HMI tags "DB_SDC_ERROR_STAT_EMS057"
   "DB_SDC_ERRORS_STAT_ER_AKT[57].ER_TRIGER" : Word = PLC DB_SDC_ERRORS_STAT.ER_AKT[57].ER_TRIGER AT %DB3724.DBW31716, 1 s
   "DB_SDC_ERRORS_STAT_ER_AKT[57].ER_STAT[1].DRIVE_POS" : DInt = PLC DB_SDC_ERRORS_STAT.ER_AKT[57].ER_STAT[1].DRIVE_POS AT %DB3724.DBD31722, 1 s
   "DB_SDC_ERRORS_STAT_ER_AKT[57].ER_STAT[1].ERROR" : Int = PLC DB_SDC_ERRORS_STAT.ER_AKT[57].ER_STAT[1].ERROR AT %DB3724.DBW31728, 1 s
   "DB_SDC_ERRORS_STAT_ER_AKT[57].ER_STAT[2].DRIVE_POS" : DInt = PLC DB_SDC_ERRORS_STAT.ER_AKT[57].ER_STAT[2].DRIVE_POS AT %DB3724.DBD31738, 1 s
   "DB_SDC_ERRORS_STAT_ER_AKT[57].ER_STAT[2].ERROR" : Int = PLC DB_SDC_ERRORS_STAT.ER_AKT[57].ER_STAT[2].ERROR AT %DB3724.DBW31744, 1 s
   "DB_SDC_ERRORS_STAT_ER_AKT[57].ER_STAT[3].DRIVE_POS" : DInt = PLC DB_SDC_ERRORS_STAT.ER_AKT[57].ER_STAT[3].DRIVE_POS AT %DB3724.DBD31754, 1 s
   "DB_SDC_ERRORS_STAT_ER_AKT[57].ER_STAT[3].ERROR" : Int = PLC DB_SDC_ERRORS_STAT.ER_AKT[57].ER_STAT[3].ERROR AT %DB3724.DBW31760, 1 s
   "DB_SDC_ERRORS_STAT_ER_AKT[57].ER_STAT[4].DRIVE_POS" : DInt = PLC DB_SDC_ERRORS_STAT.ER_AKT[57].ER_STAT[4].DRIVE_POS AT %DB3724.DBD31770, 1 s
   "DB_SDC_ERRORS_STAT_ER_AKT[57].ER_STAT[4].ERROR" : Int = PLC DB_SDC_ERRORS_STAT.ER_AKT[57].ER_STAT[4].ERROR AT %DB3724.DBW31776, 1 s

HMI tags "DB_SDC_ERROR_STAT_EMS058"
   "DB_SDC_ERRORS_STAT_ER_AKT[58].ER_TRIGER" : Word = PLC DB_SDC_ERRORS_STAT.ER_AKT[58].ER_TRIGER AT %DB3724.DBW31782, 1 s
   "DB_SDC_ERRORS_STAT_ER_AKT[58].ER_STAT[1].DRIVE_POS" : DInt = PLC DB_SDC_ERRORS_STAT.ER_AKT[58].ER_STAT[1].DRIVE_POS AT %DB3724.DBD31788, 1 s
   "DB_SDC_ERRORS_STAT_ER_AKT[58].ER_STAT[1].ERROR" : Int = PLC DB_SDC_ERRORS_STAT.ER_AKT[58].ER_STAT[1].ERROR AT %DB3724.DBW31794, 1 s
   "DB_SDC_ERRORS_STAT_ER_AKT[58].ER_STAT[2].DRIVE_POS" : DInt = PLC DB_SDC_ERRORS_STAT.ER_AKT[58].ER_STAT[2].DRIVE_POS AT %DB3724.DBD31804, 1 s
   "DB_SDC_ERRORS_STAT_ER_AKT[58].ER_STAT[2].ERROR" : Int = PLC DB_SDC_ERRORS_STAT.ER_AKT[58].ER_STAT[2].ERROR AT %DB3724.DBW31810, 1 s
   "DB_SDC_ERRORS_STAT_ER_AKT[58].ER_STAT[3].DRIVE_POS" : DInt = PLC DB_SDC_ERRORS_STAT.ER_AKT[58].ER_STAT[3].DRIVE_POS AT %DB3724.DBD31820, 1 s
   "DB_SDC_ERRORS_STAT_ER_AKT[58].ER_STAT[3].ERROR" : Int = PLC DB_SDC_ERRORS_STAT.ER_AKT[58].ER_STAT[3].ERROR AT %DB3724.DBW31826, 1 s
   "DB_SDC_ERRORS_STAT_ER_AKT[58].ER_STAT[4].DRIVE_POS" : DInt = PLC DB_SDC_ERRORS_STAT.ER_AKT[58].ER_STAT[4].DRIVE_POS AT %DB3724.DBD31836, 1 s
   "DB_SDC_ERRORS_STAT_ER_AKT[58].ER_STAT[4].ERROR" : Int = PLC DB_SDC_ERRORS_STAT.ER_AKT[58].ER_STAT[4].ERROR AT %DB3724.DBW31842, 1 s

HMI tags "DB_SDC_ERROR_STAT_EMS059"
   "DB_SDC_ERRORS_STAT_ER_AKT[59].ER_TRIGER" : Word = PLC DB_SDC_ERRORS_STAT.ER_AKT[59].ER_TRIGER AT %DB3724.DBW31848, 1 s
   "DB_SDC_ERRORS_STAT_ER_AKT[59].ER_STAT[1].DRIVE_POS" : DInt = PLC DB_SDC_ERRORS_STAT.ER_AKT[59].ER_STAT[1].DRIVE_POS AT %DB3724.DBD31854, 1 s
   "DB_SDC_ERRORS_STAT_ER_AKT[59].ER_STAT[1].ERROR" : Int = PLC DB_SDC_ERRORS_STAT.ER_AKT[59].ER_STAT[1].ERROR AT %DB3724.DBW31860, 1 s
   "DB_SDC_ERRORS_STAT_ER_AKT[59].ER_STAT[2].DRIVE_POS" : DInt = PLC DB_SDC_ERRORS_STAT.ER_AKT[59].ER_STAT[2].DRIVE_POS AT %DB3724.DBD31870, 1 s
   "DB_SDC_ERRORS_STAT_ER_AKT[59].ER_STAT[2].ERROR" : Int = PLC DB_SDC_ERRORS_STAT.ER_AKT[59].ER_STAT[2].ERROR AT %DB3724.DBW31876, 1 s
   "DB_SDC_ERRORS_STAT_ER_AKT[59].ER_STAT[3].DRIVE_POS" : DInt = PLC DB_SDC_ERRORS_STAT.ER_AKT[59].ER_STAT[3].DRIVE_POS AT %DB3724.DBD31886, 1 s
   "DB_SDC_ERRORS_STAT_ER_AKT[59].ER_STAT[3].ERROR" : Int = PLC DB_SDC_ERRORS_STAT.ER_AKT[59].ER_STAT[3].ERROR AT %DB3724.DBW31892, 1 s
   "DB_SDC_ERRORS_STAT_ER_AKT[59].ER_STAT[4].DRIVE_POS" : DInt = PLC DB_SDC_ERRORS_STAT.ER_AKT[59].ER_STAT[4].DRIVE_POS AT %DB3724.DBD31902, 1 s
   "DB_SDC_ERRORS_STAT_ER_AKT[59].ER_STAT[4].ERROR" : Int = PLC DB_SDC_ERRORS_STAT.ER_AKT[59].ER_STAT[4].ERROR AT %DB3724.DBW31908, 1 s

HMI tags "DB_SDC_ERROR_STAT_EMS060"
   "DB_SDC_ERRORS_STAT_ER_AKT[60].ER_TRIGER" : Word = PLC DB_SDC_ERRORS_STAT.ER_AKT[60].ER_TRIGER AT %DB3724.DBW31914, 1 s
   "DB_SDC_ERRORS_STAT_ER_AKT[60].ER_STAT[1].DRIVE_POS" : DInt = PLC DB_SDC_ERRORS_STAT.ER_AKT[60].ER_STAT[1].DRIVE_POS AT %DB3724.DBD31920, 1 s
   "DB_SDC_ERRORS_STAT_ER_AKT[60].ER_STAT[1].ERROR" : Int = PLC DB_SDC_ERRORS_STAT.ER_AKT[60].ER_STAT[1].ERROR AT %DB3724.DBW31926, 1 s
   "DB_SDC_ERRORS_STAT_ER_AKT[60].ER_STAT[2].DRIVE_POS" : DInt = PLC DB_SDC_ERRORS_STAT.ER_AKT[60].ER_STAT[2].DRIVE_POS AT %DB3724.DBD31936, 1 s
   "DB_SDC_ERRORS_STAT_ER_AKT[60].ER_STAT[2].ERROR" : Int = PLC DB_SDC_ERRORS_STAT.ER_AKT[60].ER_STAT[2].ERROR AT %DB3724.DBW31942, 1 s
   "DB_SDC_ERRORS_STAT_ER_AKT[60].ER_STAT[3].DRIVE_POS" : DInt = PLC DB_SDC_ERRORS_STAT.ER_AKT[60].ER_STAT[3].DRIVE_POS AT %DB3724.DBD31952, 1 s
   "DB_SDC_ERRORS_STAT_ER_AKT[60].ER_STAT[3].ERROR" : Int = PLC DB_SDC_ERRORS_STAT.ER_AKT[60].ER_STAT[3].ERROR AT %DB3724.DBW31958, 1 s
   "DB_SDC_ERRORS_STAT_ER_AKT[60].ER_STAT[4].DRIVE_POS" : DInt = PLC DB_SDC_ERRORS_STAT.ER_AKT[60].ER_STAT[4].DRIVE_POS AT %DB3724.DBD31968, 1 s
   "DB_SDC_ERRORS_STAT_ER_AKT[60].ER_STAT[4].ERROR" : Int = PLC DB_SDC_ERRORS_STAT.ER_AKT[60].ER_STAT[4].ERROR AT %DB3724.DBW31974, 1 s

HMI tags "DB_SDC_ERROR_STAT_EMS061"
   "DB_SDC_ERRORS_STAT_ER_AKT[61].ER_TRIGER" : Word = PLC DB_SDC_ERRORS_STAT.ER_AKT[61].ER_TRIGER AT %DB3724.DBW31980, 1 s
   "DB_SDC_ERRORS_STAT_ER_AKT[61].ER_STAT[1].DRIVE_POS" : DInt = PLC DB_SDC_ERRORS_STAT.ER_AKT[61].ER_STAT[1].DRIVE_POS AT %DB3724.DBD31986, 1 s
   "DB_SDC_ERRORS_STAT_ER_AKT[61].ER_STAT[1].ERROR" : Int = PLC DB_SDC_ERRORS_STAT.ER_AKT[61].ER_STAT[1].ERROR AT %DB3724.DBW31992, 1 s
   "DB_SDC_ERRORS_STAT_ER_AKT[61].ER_STAT[2].DRIVE_POS" : DInt = PLC DB_SDC_ERRORS_STAT.ER_AKT[61].ER_STAT[2].DRIVE_POS AT %DB3724.DBD32002, 1 s
   "DB_SDC_ERRORS_STAT_ER_AKT[61].ER_STAT[2].ERROR" : Int = PLC DB_SDC_ERRORS_STAT.ER_AKT[61].ER_STAT[2].ERROR AT %DB3724.DBW32008, 1 s
   "DB_SDC_ERRORS_STAT_ER_AKT[61].ER_STAT[3].DRIVE_POS" : DInt = PLC DB_SDC_ERRORS_STAT.ER_AKT[61].ER_STAT[3].DRIVE_POS AT %DB3724.DBD32018, 1 s
   "DB_SDC_ERRORS_STAT_ER_AKT[61].ER_STAT[3].ERROR" : Int = PLC DB_SDC_ERRORS_STAT.ER_AKT[61].ER_STAT[3].ERROR AT %DB3724.DBW32024, 1 s
   "DB_SDC_ERRORS_STAT_ER_AKT[61].ER_STAT[4].DRIVE_POS" : DInt = PLC DB_SDC_ERRORS_STAT.ER_AKT[61].ER_STAT[4].DRIVE_POS AT %DB3724.DBD32034, 1 s
   "DB_SDC_ERRORS_STAT_ER_AKT[61].ER_STAT[4].ERROR" : Int = PLC DB_SDC_ERRORS_STAT.ER_AKT[61].ER_STAT[4].ERROR AT %DB3724.DBW32040, 1 s

HMI tags "DB_SDC_ERROR_STAT_EMS062"
   "DB_SDC_ERRORS_STAT_ER_AKT[62].ER_TRIGER" : Word = PLC DB_SDC_ERRORS_STAT.ER_AKT[62].ER_TRIGER AT %DB3724.DBW32046, 1 s
   "DB_SDC_ERRORS_STAT_ER_AKT[62].ER_STAT[1].DRIVE_POS" : DInt = PLC DB_SDC_ERRORS_STAT.ER_AKT[62].ER_STAT[1].DRIVE_POS AT %DB3724.DBD32052, 1 s
   "DB_SDC_ERRORS_STAT_ER_AKT[62].ER_STAT[1].ERROR" : Int = PLC DB_SDC_ERRORS_STAT.ER_AKT[62].ER_STAT[1].ERROR AT %DB3724.DBW32058, 1 s
   "DB_SDC_ERRORS_STAT_ER_AKT[62].ER_STAT[2].DRIVE_POS" : DInt = PLC DB_SDC_ERRORS_STAT.ER_AKT[62].ER_STAT[2].DRIVE_POS AT %DB3724.DBD32068, 1 s
   "DB_SDC_ERRORS_STAT_ER_AKT[62].ER_STAT[2].ERROR" : Int = PLC DB_SDC_ERRORS_STAT.ER_AKT[62].ER_STAT[2].ERROR AT %DB3724.DBW32074, 1 s
   "DB_SDC_ERRORS_STAT_ER_AKT[62].ER_STAT[3].DRIVE_POS" : DInt = PLC DB_SDC_ERRORS_STAT.ER_AKT[62].ER_STAT[3].DRIVE_POS AT %DB3724.DBD32084, 1 s
   "DB_SDC_ERRORS_STAT_ER_AKT[62].ER_STAT[3].ERROR" : Int = PLC DB_SDC_ERRORS_STAT.ER_AKT[62].ER_STAT[3].ERROR AT %DB3724.DBW32090, 1 s
   "DB_SDC_ERRORS_STAT_ER_AKT[62].ER_STAT[4].DRIVE_POS" : DInt = PLC DB_SDC_ERRORS_STAT.ER_AKT[62].ER_STAT[4].DRIVE_POS AT %DB3724.DBD32100, 1 s
   "DB_SDC_ERRORS_STAT_ER_AKT[62].ER_STAT[4].ERROR" : Int = PLC DB_SDC_ERRORS_STAT.ER_AKT[62].ER_STAT[4].ERROR AT %DB3724.DBW32106, 1 s

HMI tags "DB_SDC_ERROR_STAT_EMS063"
   "DB_SDC_ERRORS_STAT_ER_AKT[63].ER_TRIGER" : Word = PLC DB_SDC_ERRORS_STAT.ER_AKT[63].ER_TRIGER AT %DB3724.DBW32112, 1 s
   "DB_SDC_ERRORS_STAT_ER_AKT[63].ER_STAT[1].DRIVE_POS" : DInt = PLC DB_SDC_ERRORS_STAT.ER_AKT[63].ER_STAT[1].DRIVE_POS AT %DB3724.DBD32118, 1 s
   "DB_SDC_ERRORS_STAT_ER_AKT[63].ER_STAT[1].ERROR" : Int = PLC DB_SDC_ERRORS_STAT.ER_AKT[63].ER_STAT[1].ERROR AT %DB3724.DBW32124, 1 s
   "DB_SDC_ERRORS_STAT_ER_AKT[63].ER_STAT[2].DRIVE_POS" : DInt = PLC DB_SDC_ERRORS_STAT.ER_AKT[63].ER_STAT[2].DRIVE_POS AT %DB3724.DBD32134, 1 s
   "DB_SDC_ERRORS_STAT_ER_AKT[63].ER_STAT[2].ERROR" : Int = PLC DB_SDC_ERRORS_STAT.ER_AKT[63].ER_STAT[2].ERROR AT %DB3724.DBW32140, 1 s
   "DB_SDC_ERRORS_STAT_ER_AKT[63].ER_STAT[3].DRIVE_POS" : DInt = PLC DB_SDC_ERRORS_STAT.ER_AKT[63].ER_STAT[3].DRIVE_POS AT %DB3724.DBD32150, 1 s
   "DB_SDC_ERRORS_STAT_ER_AKT[63].ER_STAT[3].ERROR" : Int = PLC DB_SDC_ERRORS_STAT.ER_AKT[63].ER_STAT[3].ERROR AT %DB3724.DBW32156, 1 s
   "DB_SDC_ERRORS_STAT_ER_AKT[63].ER_STAT[4].DRIVE_POS" : DInt = PLC DB_SDC_ERRORS_STAT.ER_AKT[63].ER_STAT[4].DRIVE_POS AT %DB3724.DBD32166, 1 s
   "DB_SDC_ERRORS_STAT_ER_AKT[63].ER_STAT[4].ERROR" : Int = PLC DB_SDC_ERRORS_STAT.ER_AKT[63].ER_STAT[4].ERROR AT %DB3724.DBW32172, 1 s

HMI tags "DB_SDC_ERROR_STAT_EMS064"
   "DB_SDC_ERRORS_STAT_ER_AKT[64].ER_TRIGER" : Word = PLC DB_SDC_ERRORS_STAT.ER_AKT[64].ER_TRIGER AT %DB3724.DBW32178, 1 s
   "DB_SDC_ERRORS_STAT_ER_AKT[64].ER_STAT[1].DRIVE_POS" : DInt = PLC DB_SDC_ERRORS_STAT.ER_AKT[64].ER_STAT[1].DRIVE_POS AT %DB3724.DBD32184, 1 s
   "DB_SDC_ERRORS_STAT_ER_AKT[64].ER_STAT[1].ERROR" : Int = PLC DB_SDC_ERRORS_STAT.ER_AKT[64].ER_STAT[1].ERROR AT %DB3724.DBW32190, 1 s
   "DB_SDC_ERRORS_STAT_ER_AKT[64].ER_STAT[2].DRIVE_POS" : DInt = PLC DB_SDC_ERRORS_STAT.ER_AKT[64].ER_STAT[2].DRIVE_POS AT %DB3724.DBD32200, 1 s
   "DB_SDC_ERRORS_STAT_ER_AKT[64].ER_STAT[2].ERROR" : Int = PLC DB_SDC_ERRORS_STAT.ER_AKT[64].ER_STAT[2].ERROR AT %DB3724.DBW32206, 1 s
   "DB_SDC_ERRORS_STAT_ER_AKT[64].ER_STAT[3].DRIVE_POS" : DInt = PLC DB_SDC_ERRORS_STAT.ER_AKT[64].ER_STAT[3].DRIVE_POS AT %DB3724.DBD32216, 1 s
   "DB_SDC_ERRORS_STAT_ER_AKT[64].ER_STAT[3].ERROR" : Int = PLC DB_SDC_ERRORS_STAT.ER_AKT[64].ER_STAT[3].ERROR AT %DB3724.DBW32222, 1 s
   "DB_SDC_ERRORS_STAT_ER_AKT[64].ER_STAT[4].DRIVE_POS" : DInt = PLC DB_SDC_ERRORS_STAT.ER_AKT[64].ER_STAT[4].DRIVE_POS AT %DB3724.DBD32232, 1 s
   "DB_SDC_ERRORS_STAT_ER_AKT[64].ER_STAT[4].ERROR" : Int = PLC DB_SDC_ERRORS_STAT.ER_AKT[64].ER_STAT[4].ERROR AT %DB3724.DBW32238, 1 s

HMI tags "DB_SDC_ERROR_STAT_EMS065"
   "DB_SDC_ERRORS_STAT_ER_AKT[65].ER_TRIGER" : Word = PLC DB_SDC_ERRORS_STAT.ER_AKT[65].ER_TRIGER AT %DB3724.DBW32244, 1 s
   "DB_SDC_ERRORS_STAT_ER_AKT[65].ER_STAT[1].DRIVE_POS" : DInt = PLC DB_SDC_ERRORS_STAT.ER_AKT[65].ER_STAT[1].DRIVE_POS AT %DB3724.DBD32250, 1 s
   "DB_SDC_ERRORS_STAT_ER_AKT[65].ER_STAT[1].ERROR" : Int = PLC DB_SDC_ERRORS_STAT.ER_AKT[65].ER_STAT[1].ERROR AT %DB3724.DBW32256, 1 s
   "DB_SDC_ERRORS_STAT_ER_AKT[65].ER_STAT[2].DRIVE_POS" : DInt = PLC DB_SDC_ERRORS_STAT.ER_AKT[65].ER_STAT[2].DRIVE_POS AT %DB3724.DBD32266, 1 s
   "DB_SDC_ERRORS_STAT_ER_AKT[65].ER_STAT[2].ERROR" : Int = PLC DB_SDC_ERRORS_STAT.ER_AKT[65].ER_STAT[2].ERROR AT %DB3724.DBW32272, 1 s
   "DB_SDC_ERRORS_STAT_ER_AKT[65].ER_STAT[3].DRIVE_POS" : DInt = PLC DB_SDC_ERRORS_STAT.ER_AKT[65].ER_STAT[3].DRIVE_POS AT %DB3724.DBD32282, 1 s
   "DB_SDC_ERRORS_STAT_ER_AKT[65].ER_STAT[3].ERROR" : Int = PLC DB_SDC_ERRORS_STAT.ER_AKT[65].ER_STAT[3].ERROR AT %DB3724.DBW32288, 1 s
   "DB_SDC_ERRORS_STAT_ER_AKT[65].ER_STAT[4].DRIVE_POS" : DInt = PLC DB_SDC_ERRORS_STAT.ER_AKT[65].ER_STAT[4].DRIVE_POS AT %DB3724.DBD32298, 1 s
   "DB_SDC_ERRORS_STAT_ER_AKT[65].ER_STAT[4].ERROR" : Int = PLC DB_SDC_ERRORS_STAT.ER_AKT[65].ER_STAT[4].ERROR AT %DB3724.DBW32304, 1 s

HMI tags "DB_SDC_ERROR_STAT_EMS066"
   "DB_SDC_ERRORS_STAT_ER_AKT[66].ER_TRIGER" : Word = PLC DB_SDC_ERRORS_STAT.ER_AKT[66].ER_TRIGER AT %DB3724.DBW32310, 1 s
   "DB_SDC_ERRORS_STAT_ER_AKT[66].ER_STAT[1].DRIVE_POS" : DInt = PLC DB_SDC_ERRORS_STAT.ER_AKT[66].ER_STAT[1].DRIVE_POS AT %DB3724.DBD32316, 1 s
   "DB_SDC_ERRORS_STAT_ER_AKT[66].ER_STAT[1].ERROR" : Int = PLC DB_SDC_ERRORS_STAT.ER_AKT[66].ER_STAT[1].ERROR AT %DB3724.DBW32322, 1 s
   "DB_SDC_ERRORS_STAT_ER_AKT[66].ER_STAT[2].DRIVE_POS" : DInt = PLC DB_SDC_ERRORS_STAT.ER_AKT[66].ER_STAT[2].DRIVE_POS AT %DB3724.DBD32332, 1 s
   "DB_SDC_ERRORS_STAT_ER_AKT[66].ER_STAT[2].ERROR" : Int = PLC DB_SDC_ERRORS_STAT.ER_AKT[66].ER_STAT[2].ERROR AT %DB3724.DBW32338, 1 s
   "DB_SDC_ERRORS_STAT_ER_AKT[66].ER_STAT[3].DRIVE_POS" : DInt = PLC DB_SDC_ERRORS_STAT.ER_AKT[66].ER_STAT[3].DRIVE_POS AT %DB3724.DBD32348, 1 s
   "DB_SDC_ERRORS_STAT_ER_AKT[66].ER_STAT[3].ERROR" : Int = PLC DB_SDC_ERRORS_STAT.ER_AKT[66].ER_STAT[3].ERROR AT %DB3724.DBW32354, 1 s
   "DB_SDC_ERRORS_STAT_ER_AKT[66].ER_STAT[4].DRIVE_POS" : DInt = PLC DB_SDC_ERRORS_STAT.ER_AKT[66].ER_STAT[4].DRIVE_POS AT %DB3724.DBD32364, 1 s
   "DB_SDC_ERRORS_STAT_ER_AKT[66].ER_STAT[4].ERROR" : Int = PLC DB_SDC_ERRORS_STAT.ER_AKT[66].ER_STAT[4].ERROR AT %DB3724.DBW32370, 1 s

HMI tags "DB_SDC_ERROR_STAT_EMS067"
   "DB_SDC_ERRORS_STAT_ER_AKT[67].ER_TRIGER" : Word = PLC DB_SDC_ERRORS_STAT.ER_AKT[67].ER_TRIGER AT %DB3724.DBW32376, 1 s
   "DB_SDC_ERRORS_STAT_ER_AKT[67].ER_STAT[1].DRIVE_POS" : DInt = PLC DB_SDC_ERRORS_STAT.ER_AKT[67].ER_STAT[1].DRIVE_POS AT %DB3724.DBD32382, 1 s
   "DB_SDC_ERRORS_STAT_ER_AKT[67].ER_STAT[1].ERROR" : Int = PLC DB_SDC_ERRORS_STAT.ER_AKT[67].ER_STAT[1].ERROR AT %DB3724.DBW32388, 1 s
   "DB_SDC_ERRORS_STAT_ER_AKT[67].ER_STAT[2].DRIVE_POS" : DInt = PLC DB_SDC_ERRORS_STAT.ER_AKT[67].ER_STAT[2].DRIVE_POS AT %DB3724.DBD32398, 1 s
   "DB_SDC_ERRORS_STAT_ER_AKT[67].ER_STAT[2].ERROR" : Int = PLC DB_SDC_ERRORS_STAT.ER_AKT[67].ER_STAT[2].ERROR AT %DB3724.DBW32404, 1 s
   "DB_SDC_ERRORS_STAT_ER_AKT[67].ER_STAT[3].DRIVE_POS" : DInt = PLC DB_SDC_ERRORS_STAT.ER_AKT[67].ER_STAT[3].DRIVE_POS AT %DB3724.DBD32414, 1 s
   "DB_SDC_ERRORS_STAT_ER_AKT[67].ER_STAT[3].ERROR" : Int = PLC DB_SDC_ERRORS_STAT.ER_AKT[67].ER_STAT[3].ERROR AT %DB3724.DBW32420, 1 s
   "DB_SDC_ERRORS_STAT_ER_AKT[67].ER_STAT[4].DRIVE_POS" : DInt = PLC DB_SDC_ERRORS_STAT.ER_AKT[67].ER_STAT[4].DRIVE_POS AT %DB3724.DBD32430, 1 s
   "DB_SDC_ERRORS_STAT_ER_AKT[67].ER_STAT[4].ERROR" : Int = PLC DB_SDC_ERRORS_STAT.ER_AKT[67].ER_STAT[4].ERROR AT %DB3724.DBW32436, 1 s

HMI tags "DB_SDC_ERROR_STAT_EMS068"
   "DB_SDC_ERRORS_STAT_ER_AKT[68].ER_TRIGER" : Word = PLC DB_SDC_ERRORS_STAT.ER_AKT[68].ER_TRIGER AT %DB3724.DBW32442, 1 s
   "DB_SDC_ERRORS_STAT_ER_AKT[68].ER_STAT[1].DRIVE_POS" : DInt = PLC DB_SDC_ERRORS_STAT.ER_AKT[68].ER_STAT[1].DRIVE_POS AT %DB3724.DBD32448, 1 s
   "DB_SDC_ERRORS_STAT_ER_AKT[68].ER_STAT[1].ERROR" : Int = PLC DB_SDC_ERRORS_STAT.ER_AKT[68].ER_STAT[1].ERROR AT %DB3724.DBW32454, 1 s
   "DB_SDC_ERRORS_STAT_ER_AKT[68].ER_STAT[2].DRIVE_POS" : DInt = PLC DB_SDC_ERRORS_STAT.ER_AKT[68].ER_STAT[2].DRIVE_POS AT %DB3724.DBD32464, 1 s
   "DB_SDC_ERRORS_STAT_ER_AKT[68].ER_STAT[2].ERROR" : Int = PLC DB_SDC_ERRORS_STAT.ER_AKT[68].ER_STAT[2].ERROR AT %DB3724.DBW32470, 1 s
   "DB_SDC_ERRORS_STAT_ER_AKT[68].ER_STAT[3].DRIVE_POS" : DInt = PLC DB_SDC_ERRORS_STAT.ER_AKT[68].ER_STAT[3].DRIVE_POS AT %DB3724.DBD32480, 1 s
   "DB_SDC_ERRORS_STAT_ER_AKT[68].ER_STAT[3].ERROR" : Int = PLC DB_SDC_ERRORS_STAT.ER_AKT[68].ER_STAT[3].ERROR AT %DB3724.DBW32486, 1 s
   "DB_SDC_ERRORS_STAT_ER_AKT[68].ER_STAT[4].DRIVE_POS" : DInt = PLC DB_SDC_ERRORS_STAT.ER_AKT[68].ER_STAT[4].DRIVE_POS AT %DB3724.DBD32496, 1 s
   "DB_SDC_ERRORS_STAT_ER_AKT[68].ER_STAT[4].ERROR" : Int = PLC DB_SDC_ERRORS_STAT.ER_AKT[68].ER_STAT[4].ERROR AT %DB3724.DBW32502, 1 s

HMI tags "DB_SDC_ERROR_STAT_EMS069"
   "DB_SDC_ERRORS_STAT_ER_AKT[69].ER_TRIGER" : Word = PLC DB_SDC_ERRORS_STAT.ER_AKT[69].ER_TRIGER AT %DB3724.DBW32508, 1 s
   "DB_SDC_ERRORS_STAT_ER_AKT[69].ER_STAT[1].DRIVE_POS" : DInt = PLC DB_SDC_ERRORS_STAT.ER_AKT[69].ER_STAT[1].DRIVE_POS AT %DB3724.DBD32514, 1 s
   "DB_SDC_ERRORS_STAT_ER_AKT[69].ER_STAT[1].ERROR" : Int = PLC DB_SDC_ERRORS_STAT.ER_AKT[69].ER_STAT[1].ERROR AT %DB3724.DBW32520, 1 s
   "DB_SDC_ERRORS_STAT_ER_AKT[69].ER_STAT[2].DRIVE_POS" : DInt = PLC DB_SDC_ERRORS_STAT.ER_AKT[69].ER_STAT[2].DRIVE_POS AT %DB3724.DBD32530, 1 s
   "DB_SDC_ERRORS_STAT_ER_AKT[69].ER_STAT[2].ERROR" : Int = PLC DB_SDC_ERRORS_STAT.ER_AKT[69].ER_STAT[2].ERROR AT %DB3724.DBW32536, 1 s
   "DB_SDC_ERRORS_STAT_ER_AKT[69].ER_STAT[3].DRIVE_POS" : DInt = PLC DB_SDC_ERRORS_STAT.ER_AKT[69].ER_STAT[3].DRIVE_POS AT %DB3724.DBD32546, 1 s
   "DB_SDC_ERRORS_STAT_ER_AKT[69].ER_STAT[3].ERROR" : Int = PLC DB_SDC_ERRORS_STAT.ER_AKT[69].ER_STAT[3].ERROR AT %DB3724.DBW32552, 1 s
   "DB_SDC_ERRORS_STAT_ER_AKT[69].ER_STAT[4].DRIVE_POS" : DInt = PLC DB_SDC_ERRORS_STAT.ER_AKT[69].ER_STAT[4].DRIVE_POS AT %DB3724.DBD32562, 1 s
   "DB_SDC_ERRORS_STAT_ER_AKT[69].ER_STAT[4].ERROR" : Int = PLC DB_SDC_ERRORS_STAT.ER_AKT[69].ER_STAT[4].ERROR AT %DB3724.DBW32568, 1 s

HMI tags "DB_SDC_ERROR_STAT_EMS070"
   "DB_SDC_ERRORS_STAT_ER_AKT[70].ER_TRIGER" : Word = PLC DB_SDC_ERRORS_STAT.ER_AKT[70].ER_TRIGER AT %DB3724.DBW32574, 1 s
   "DB_SDC_ERRORS_STAT_ER_AKT[70].ER_STAT[1].DRIVE_POS" : DInt = PLC DB_SDC_ERRORS_STAT.ER_AKT[70].ER_STAT[1].DRIVE_POS AT %DB3724.DBD32580, 1 s
   "DB_SDC_ERRORS_STAT_ER_AKT[70].ER_STAT[1].ERROR" : Int = PLC DB_SDC_ERRORS_STAT.ER_AKT[70].ER_STAT[1].ERROR AT %DB3724.DBW32586, 1 s
   "DB_SDC_ERRORS_STAT_ER_AKT[70].ER_STAT[2].DRIVE_POS" : DInt = PLC DB_SDC_ERRORS_STAT.ER_AKT[70].ER_STAT[2].DRIVE_POS AT %DB3724.DBD32596, 1 s
   "DB_SDC_ERRORS_STAT_ER_AKT[70].ER_STAT[2].ERROR" : Int = PLC DB_SDC_ERRORS_STAT.ER_AKT[70].ER_STAT[2].ERROR AT %DB3724.DBW32602, 1 s
   "DB_SDC_ERRORS_STAT_ER_AKT[70].ER_STAT[3].DRIVE_POS" : DInt = PLC DB_SDC_ERRORS_STAT.ER_AKT[70].ER_STAT[3].DRIVE_POS AT %DB3724.DBD32612, 1 s
   "DB_SDC_ERRORS_STAT_ER_AKT[70].ER_STAT[3].ERROR" : Int = PLC DB_SDC_ERRORS_STAT.ER_AKT[70].ER_STAT[3].ERROR AT %DB3724.DBW32618, 1 s
   "DB_SDC_ERRORS_STAT_ER_AKT[70].ER_STAT[4].DRIVE_POS" : DInt = PLC DB_SDC_ERRORS_STAT.ER_AKT[70].ER_STAT[4].DRIVE_POS AT %DB3724.DBD32628, 1 s
   "DB_SDC_ERRORS_STAT_ER_AKT[70].ER_STAT[4].ERROR" : Int = PLC DB_SDC_ERRORS_STAT.ER_AKT[70].ER_STAT[4].ERROR AT %DB3724.DBW32634, 1 s

HMI tags "DB_SDC_ERROR_STAT_EMS071"
   "DB_SDC_ERRORS_STAT_ER_AKT[71].ER_TRIGER" : Word = PLC DB_SDC_ERRORS_STAT.ER_AKT[71].ER_TRIGER AT %DB3724.DBW32640, 1 s
   "DB_SDC_ERRORS_STAT_ER_AKT[71].ER_STAT[1].DRIVE_POS" : DInt = PLC DB_SDC_ERRORS_STAT.ER_AKT[71].ER_STAT[1].DRIVE_POS AT %DB3724.DBD32646, 1 s
   "DB_SDC_ERRORS_STAT_ER_AKT[71].ER_STAT[1].ERROR" : Int = PLC DB_SDC_ERRORS_STAT.ER_AKT[71].ER_STAT[1].ERROR AT %DB3724.DBW32652, 1 s
   "DB_SDC_ERRORS_STAT_ER_AKT[71].ER_STAT[2].DRIVE_POS" : DInt = PLC DB_SDC_ERRORS_STAT.ER_AKT[71].ER_STAT[2].DRIVE_POS AT %DB3724.DBD32662, 1 s
   "DB_SDC_ERRORS_STAT_ER_AKT[71].ER_STAT[2].ERROR" : Int = PLC DB_SDC_ERRORS_STAT.ER_AKT[71].ER_STAT[2].ERROR AT %DB3724.DBW32668, 1 s
   "DB_SDC_ERRORS_STAT_ER_AKT[71].ER_STAT[3].DRIVE_POS" : DInt = PLC DB_SDC_ERRORS_STAT.ER_AKT[71].ER_STAT[3].DRIVE_POS AT %DB3724.DBD32678, 1 s
   "DB_SDC_ERRORS_STAT_ER_AKT[71].ER_STAT[3].ERROR" : Int = PLC DB_SDC_ERRORS_STAT.ER_AKT[71].ER_STAT[3].ERROR AT %DB3724.DBW32684, 1 s
   "DB_SDC_ERRORS_STAT_ER_AKT[71].ER_STAT[4].DRIVE_POS" : DInt = PLC DB_SDC_ERRORS_STAT.ER_AKT[71].ER_STAT[4].DRIVE_POS AT %DB3724.DBD32694, 1 s
   "DB_SDC_ERRORS_STAT_ER_AKT[71].ER_STAT[4].ERROR" : Int = PLC DB_SDC_ERRORS_STAT.ER_AKT[71].ER_STAT[4].ERROR AT %DB3724.DBW32700, 1 s

HMI tags "DB_SDC_ERROR_STAT_EMS072"
   "DB_SDC_ERRORS_STAT_ER_AKT[72].ER_TRIGER" : Word = PLC DB_SDC_ERRORS_STAT.ER_AKT[72].ER_TRIGER AT %DB3724.DBW32706, 1 s
   "DB_SDC_ERRORS_STAT_ER_AKT[72].ER_STAT[1].DRIVE_POS" : DInt = PLC DB_SDC_ERRORS_STAT.ER_AKT[72].ER_STAT[1].DRIVE_POS AT %DB3724.DBD32712, 1 s
   "DB_SDC_ERRORS_STAT_ER_AKT[72].ER_STAT[1].ERROR" : Int = PLC DB_SDC_ERRORS_STAT.ER_AKT[72].ER_STAT[1].ERROR AT %DB3724.DBW32718, 1 s
   "DB_SDC_ERRORS_STAT_ER_AKT[72].ER_STAT[2].DRIVE_POS" : DInt = PLC DB_SDC_ERRORS_STAT.ER_AKT[72].ER_STAT[2].DRIVE_POS AT %DB3724.DBD32728, 1 s
   "DB_SDC_ERRORS_STAT_ER_AKT[72].ER_STAT[2].ERROR" : Int = PLC DB_SDC_ERRORS_STAT.ER_AKT[72].ER_STAT[2].ERROR AT %DB3724.DBW32734, 1 s
   "DB_SDC_ERRORS_STAT_ER_AKT[72].ER_STAT[3].DRIVE_POS" : DInt = PLC DB_SDC_ERRORS_STAT.ER_AKT[72].ER_STAT[3].DRIVE_POS AT %DB3724.DBD32744, 1 s
   "DB_SDC_ERRORS_STAT_ER_AKT[72].ER_STAT[3].ERROR" : Int = PLC DB_SDC_ERRORS_STAT.ER_AKT[72].ER_STAT[3].ERROR AT %DB3724.DBW32750, 1 s
   "DB_SDC_ERRORS_STAT_ER_AKT[72].ER_STAT[4].DRIVE_POS" : DInt = PLC DB_SDC_ERRORS_STAT.ER_AKT[72].ER_STAT[4].DRIVE_POS AT %DB3724.DBD32760, 1 s
   "DB_SDC_ERRORS_STAT_ER_AKT[72].ER_STAT[4].ERROR" : Int = PLC DB_SDC_ERRORS_STAT.ER_AKT[72].ER_STAT[4].ERROR AT %DB3724.DBW32766, 1 s

HMI tags "VAT_DB_SDC_EMS_FLAGS"
   "SDC\DB_SDC_EMS_FLAGS\DB_SDC_EMS_FLAGS.EMS[8]" : Int AT %DB0.DBW0, 1 s   // EMSdriver present
   "SDC\DB_SDC_EMS_FLAGS\_EMS_Flags_HMI_Byte_00" : Int, internal
   "SDC\DB_SDC_EMS_FLAGS\_EMS_Flags_HMI_Byte_19" : Int, internal
   "DB_SDC_EMS_FLAGS_HMI_HMI[1].RET_VAL_SFC12" : Int = PLC DB_SDC_EMS_FLAGS_HMI.HMI[1].RET_VAL_SFC12 AT %DB3801.DBW34, 1 s   // RetVal SFC12
   "SDC\DB_SDC_EMS_FLAGS\DB_SDC_EMS_FLAGS.EMS[9]" : Int AT %DB0.DBW0, 1 s   // EMSdriver present
   "SDC\DB_SDC_EMS_FLAGS\DB_SDC_EMS_FLAGS.EMS[19]" : Int AT %DB0.DBW0, 1 s   // EMSdriver present
   "SDC\DB_SDC_EMS_FLAGS\DB_SDC_EMS_FLAGS.HMI[XX].EMS_Nr" : Int AT %DB0.DBW0, 1 s   // Sektionsnummer
   "SDC\DB_SDC_EMS_FLAGS\_EMS_Flags_HMI_Byte_04" : Int, internal
   "SDC\DB_SDC_EMS_FLAGS\DB_SDC_EMS_FLAGS.HMI[XX].PULT_Nr_EDIT" : Int AT %DB0.DBW0, 1 s   // Pult Nr Editieren Aktiv (HMI 1 = Master)
   "SDC\DB_SDC_EMS_FLAGS\DB_SDC_EMS_FLAGS.EMS[20]" : Int AT %DB0.DBW0, 1 s   // EMSdriver present
   "DB_SDC_EMS_FLAGS_HEADER.LAENGE_EMS_FLAGS" : Int = PLC DB_SDC_EMS_FLAGS.HEADER.LAENGE_EMS_FLAGS AT %DB3701.DBW8, 1 s   // Länge Eingänge pro EMS
   "SDC\DB_SDC_EMS_FLAGS\DB_SDC_EMS_FLAGS.EMS[6]" : Int AT %DB0.DBW0, 1 s   // EMSdriver present
   "SDC\DB_SDC_EMS_FLAGS\DB_SDC_EMS_FLAGS.EMS[12]" : Int AT %DB0.DBW0, 1 s   // EMSdriver present
   "SDC\DB_SDC_EMS_FLAGS\DB_SDC_EMS_FLAGS.EMS[1]" : Int AT %DB0.DBW0, 1 s   // EMSdriver present
   "SDC\DB_SDC_EMS_FLAGS\DB_SDC_EMS_FLAGS.EMS[3]" : Int AT %DB0.DBW0, 1 s   // EMSdriver present
   "SDC\DB_SDC_EMS_FLAGS\DB_SDC_EMS_FLAGS.HMI[XX].BILD_Nr" : Int AT %DB0.DBW0, 1 s   // Bild_Nr aktiv
   "SDC\DB_SDC_EMS_FLAGS\DB_SDC_EMS_FLAGS.HMI[XX].T_LOAD" : Bool AT %DB0.DBX0.3, 1 s   // Taster laden
   "DB_SDC_EMS_FLAGS_HMI_HEADER.START_HMI" : Int = PLC DB_SDC_EMS_FLAGS_HMI.HEADER.START_HMI AT %DB3801.DBW10, 1 s   // Startadresse HMI
   "SDC\DB_SDC_EMS_FLAGS\DB_SDC_EMS_FLAGS.EMS[10]" : Int AT %DB0.DBW0, 1 s   // EMSdriver present
   "SDC\DB_SDC_EMS_FLAGS\_EMS_Flags_HMI_Byte_18" : Int, internal
   "SDC\DB_SDC_EMS_FLAGS\DB_SDC_EMS_FLAGS.EMS[7]" : Int AT %DB0.DBW0, 1 s   // EMSdriver present
   "SDC\DB_SDC_EMS_FLAGS\DB_SDC_EMS_FLAGS.EMS[13]" : Int AT %DB0.DBW0, 1 s   // EMSdriver present
   "DB_SDC_EMS_FLAGS_HMI_HMI[1].MODE_SFC12" : Byte = PLC DB_SDC_EMS_FLAGS_HMI.HMI[1].MODE_SFC12 AT %DB3801.DBB36, 1 s   // Mode SFC12
   "SDC\DB_SDC_EMS_FLAGS\DB_SDC_EMS_FLAGS.HMI[XX].FR_EDIT" : Bool AT %DB0.DBX0.0, 1 s   // Freigabe Editieren
   "SDC\DB_SDC_EMS_FLAGS\_EMS_Flags_HMI_Byte_12" : Int, internal
   "SDC\DB_SDC_EMS_FLAGS\DB_SDC_EMS_FLAGS.EMS[18]" : Int AT %DB0.DBW0, 1 s   // EMSdriver present
   "DB_SDC_EMS_FLAGS_HEADER.DB_NR" : Int = PLC DB_SDC_EMS_FLAGS.HEADER.DB_NR AT %DB3701.DBW0, 1 s   // DB Nummer
   "SDC\DB_SDC_EMS_FLAGS\DB_SDC_EMS_FLAGS.HMI[XX].BILD_Nr_Alt" : Int AT %DB0.DBW0, 1 s   // Bild_Nr alt
   "DB_SDC_EMS_FLAGS_HMI_HEADER.OFFEST_HMI_DATA" : Int = PLC DB_SDC_EMS_FLAGS_HMI.HEADER.OFFEST_HMI_DATA AT %DB3801.DBW12, 1 s   // Offestadresse der HMI Flag Data
   "SDC\DB_SDC_EMS_FLAGS\DB_SDC_EMS_FLAGS.EMS[2]" : Int AT %DB0.DBW0, 1 s   // EMSdriver present
   "DB_SDC_EMS_FLAGS_HEADER.MIN_NR_EMS" : Int = PLC DB_SDC_EMS_FLAGS.HEADER.MIN_NR_EMS AT %DB3701.DBW2, 1 s   // Niedrigste EMS Nummer im Daten DB
   "SDC\DB_SDC_EMS_FLAGS\DB_SDC_EMS_FLAGS.HMI[XX].T_ACTIV" : Bool AT %DB0.DBX0.4, 1 s   // Taster activieren
   "SDC\DB_SDC_EMS_FLAGS\DB_SDC_EMS_FLAGS.EMS[16]" : Int AT %DB0.DBW0, 1 s   // EMSdriver present
   "SDC\DB_SDC_EMS_FLAGS\DB_SDC_EMS_FLAGS.HMI[XX].T_DEACTIV" : Bool AT %DB0.DBX0.5, 1 s   // Taster deactivieren
   "DB_SDC_EMS_FLAGS_HEADER.MAX_NR_EMS" : Int = PLC DB_SDC_EMS_FLAGS.HEADER.MAX_NR_EMS AT %DB3701.DBW4, 1 s   // Höchste EMS Nummer im Daten DB
   "DB_SDC_EMS_FLAGS_HMI_HMI[1].REQ_SFC12" : Bool = PLC DB_SDC_EMS_FLAGS_HMI.HMI[1].REQ_SFC12 AT %DB3801.DBX39.3, 1 s   // Request SFC12
   "SDC\DB_SDC_EMS_FLAGS\DB_SDC_EMS_FLAGS.HMI[XX].T_RESET_BED" : Bool AT %DB0.DBX0.1, 1 s   // Taster Reset Bedienfreigabe Pult Nr Bedienung
   "SDC\DB_SDC_EMS_FLAGS\_EMS_Flags_HMI_Byte_20" : Int, internal
   "DB_SDC_EMS_FLAGS_HMI_HMI[1].PULT_Nr_EDIT" : Int = PLC DB_SDC_EMS_FLAGS_HMI.HMI[1].PULT_Nr_EDIT AT %DB3801.DBW20, 1 s   // Pult Nr Editieren Aktiv (HMI 1 = Master)
   "SDC\DB_SDC_EMS_FLAGS\DB_SDC_EMS_FLAGS.HMI[XX].ER_DATA" : Bool AT %DB0.DBX0.1, 1 s   // Daten Fehlerhaft
   "SDC\DB_SDC_EMS_FLAGS\_EMS_Flags_HMI_Byte_08" : Int, internal
   "SDC\DB_SDC_EMS_FLAGS\DB_SDC_EMS_FLAGS.EMS[11]" : Int AT %DB0.DBW0, 1 s   // EMSdriver present
   "DB_SDC_EMS_FLAGS_HMI_HMI[1].TIME_SFC12" : Int = PLC DB_SDC_EMS_FLAGS_HMI.HMI[1].TIME_SFC12 AT %DB3801.DBW30, 1 s   // Actuelle Zeit Activieren/Deactivieren
   "SDC\DB_SDC_EMS_FLAGS\DB_SDC_EMS_FLAGS.EMS[14]" : Int AT %DB0.DBW0, 1 s   // EMSdriver present
   "SDC\DB_SDC_EMS_FLAGS\_EMS_Flags_HMI_Byte_16" : Int, internal
   "SDC\DB_SDC_EMS_FLAGS\DB_SDC_EMS_FLAGS.HMI[XX].T_SAVE" : Bool AT %DB0.DBX0.2, 1 s   // Taster speichern
   "SDC\DB_SDC_EMS_FLAGS\DB_SDC_EMS_FLAGS.EMS[15]" : Int AT %DB0.DBW0, 1 s   // EMSdriver present
   "SDC\DB_SDC_EMS_FLAGS\_EMS_Flags_HMI_Byte_10" : Int, internal
   "SDC\DB_SDC_EMS_FLAGS\_EMS_Flags_HMI_Byte_14" : Int, internal
   "SDC\DB_SDC_EMS_FLAGS\DB_SDC_EMS_FLAGS.HMI[XX].T_EDIT" : Bool AT %DB0.DBX0.0, 1 s   // Taster Editieren für Pult aktivieren
   "SDC\DB_SDC_EMS_FLAGS\_EMS_Flags_HMI_Byte_09" : Int, internal
   "DB_SDC_EMS_FLAGS_HMI_HMI[1].BUSY_SFC12" : Bool = PLC DB_SDC_EMS_FLAGS_HMI.HMI[1].BUSY_SFC12 AT %DB3801.DBX39.2, 1 s   // Busy SFC12
   "SDC\DB_SDC_EMS_FLAGS\_EMS_Nr" : Int, internal
      on ChangeValue: "SDC_TS_PARAMETER"(); "SDC_TS_REFERENCE"("SDC\DB_SDC_EMS_FLAGS\_EMS_Nr")
   "SDC\DB_SDC_EMS_FLAGS\DB_SDC_EMS_FLAGS.EMS[17]" : Int AT %DB0.DBW0, 1 s   // EMSdriver present
   "SDC\DB_SDC_EMS_FLAGS\_EMS_Flags_HMI_Byte_06" : Int, internal
   "SDC\DB_SDC_EMS_FLAGS\DB_SDC_EMS_FLAGS.HMI[XX].FLAGS" : Word AT %DB0.DBW0, 1 s   // Freigabe Editieren
   "SDC\DB_SDC_EMS_FLAGS\_EMS_Flags_HMI_Byte_02" : Int, internal
   "SDC\DB_SDC_EMS_FLAGS\DB_SDC_EMS_FLAGS.EMS[5]" : Int AT %DB0.DBW0, 1 s   // EMSdriver present
   "DB_SDC_EMS_FLAGS_HEADER.START_EMS" : Int = PLC DB_SDC_EMS_FLAGS.HEADER.START_EMS AT %DB3701.DBW6, 1 s   // Startadresse der EMS Daten im Daten DB
   "SDC\DB_SDC_EMS_FLAGS\DB_SDC_EMS_FLAGS.EMS[4]" : Int AT %DB0.DBW0, 1 s   // EMSdriver present
   "SDC\DB_SDC_EMS_FLAGS\DB_SDC_EMS_FLAGS.HMI[1].LADDR_SFC12" : Int AT %DB0.DBW32, 1 s   // Actuelle LADDR
   "SDC\DB_SDC_EMS_FLAGS\DB_SDC_EMS_FLAGS.EMS[21]" : Int AT %DB0.DBW0, 1 s   // EMSdriver present
   "SDC\DB_SDC_EMS_FLAGS\DB_SDC_EMS_FLAGS.EMS[22]" : Int AT %DB0.DBW0, 1 s
   "SDC\DB_SDC_EMS_FLAGS\DB_SDC_EMS_FLAGS.EMS[23]" : Int AT %DB0.DBW0, 1 s
   "SDC\DB_SDC_EMS_FLAGS\DB_SDC_EMS_FLAGS.EMS[24]" : Int AT %DB0.DBW0, 1 s
   "SDC\DB_SDC_EMS_FLAGS\DB_SDC_EMS_FLAGS.EMS[25]" : Int AT %DB0.DBW0, 1 s
   "SDC\DB_SDC_EMS_FLAGS\DB_SDC_EMS_FLAGS.EMS[26]" : Int AT %DB0.DBW0, 1 s
   "SDC\DB_SDC_EMS_FLAGS\DB_SDC_EMS_FLAGS.EMS[27]" : Int AT %DB0.DBW0, 1 s
   "SDC\DB_SDC_EMS_FLAGS\DB_SDC_EMS_FLAGS.EMS[28]" : Int AT %DB0.DBW0, 1 s
   "SDC\DB_SDC_EMS_FLAGS\DB_SDC_EMS_FLAGS.EMS[29]" : Int AT %DB0.DBW0, 1 s
   "SDC\DB_SDC_EMS_FLAGS\DB_SDC_EMS_FLAGS.EMS[30]" : Int AT %DB0.DBW0, 1 s
   "SDC\DB_SDC_EMS_FLAGS\DB_SDC_EMS_FLAGS.EMS[31]" : Int AT %DB0.DBW0, 1 s
   "SDC\DB_SDC_EMS_FLAGS\DB_SDC_EMS_FLAGS.EMS[32]" : Int AT %DB0.DBW0, 1 s
   "SDC\DB_SDC_EMS_FLAGS\DB_SDC_EMS_FLAGS.EMS[33]" : Int AT %DB0.DBW0, 1 s
   "SDC\DB_SDC_EMS_FLAGS\DB_SDC_EMS_FLAGS.EMS[34]" : Int AT %DB0.DBW0, 1 s
   "SDC\DB_SDC_EMS_FLAGS\DB_SDC_EMS_FLAGS.EMS[35]" : Int AT %DB0.DBW0, 1 s
   "SDC\DB_SDC_EMS_FLAGS\DB_SDC_EMS_FLAGS.EMS[36]" : Int AT %DB0.DBW0, 1 s
   "SDC\DB_SDC_EMS_FLAGS\DB_SDC_EMS_FLAGS.EMS[37]" : Int AT %DB0.DBW0, 1 s
   "SDC\DB_SDC_EMS_FLAGS\DB_SDC_EMS_FLAGS.EMS[38]" : Int AT %DB0.DBW0, 1 s
   "SDC\DB_SDC_EMS_FLAGS\DB_SDC_EMS_FLAGS.EMS[39]" : Int AT %DB0.DBW0, 1 s
   "SDC\DB_SDC_EMS_FLAGS\DB_SDC_EMS_FLAGS.EMS[40]" : Int AT %DB0.DBW0, 1 s
   "SDC\DB_SDC_EMS_FLAGS\DB_SDC_EMS_FLAGS.EMS[41]" : Int AT %DB0.DBW0, 1 s
   "SDC\DB_SDC_EMS_FLAGS\DB_SDC_EMS_FLAGS.EMS[42]" : Int AT %DB0.DBW0, 1 s
   "SDC\DB_SDC_EMS_FLAGS\DB_SDC_EMS_FLAGS.EMS[43]" : Int AT %DB0.DBW0, 1 s
   "SDC\DB_SDC_EMS_FLAGS\DB_SDC_EMS_FLAGS.EMS[44]" : Int AT %DB0.DBW0, 1 s
   "SDC\DB_SDC_EMS_FLAGS\DB_SDC_EMS_FLAGS.EMS[45]" : Int AT %DB0.DBW0, 1 s
   "SDC\DB_SDC_EMS_FLAGS\DB_SDC_EMS_FLAGS.EMS[46]" : Int AT %DB0.DBW0, 1 s
   "SDC\DB_SDC_EMS_FLAGS\DB_SDC_EMS_FLAGS.EMS[47]" : Int AT %DB0.DBW0, 1 s
   "SDC\DB_SDC_EMS_FLAGS\DB_SDC_EMS_FLAGS.EMS[48]" : Int AT %DB0.DBW0, 1 s
   "SDC\DB_SDC_EMS_FLAGS\DB_SDC_EMS_FLAGS.EMS[49]" : Int AT %DB0.DBW0, 1 s
   "SDC\DB_SDC_EMS_FLAGS\DB_SDC_EMS_FLAGS.EMS[50]" : Int AT %DB0.DBW0, 1 s
   "SDC\DB_SDC_EMS_FLAGS\DB_SDC_EMS_FLAGS.EMS[51]" : Int AT %DB0.DBW0, 1 s
   "SDC\DB_SDC_EMS_FLAGS\DB_SDC_EMS_FLAGS.EMS[52]" : Int AT %DB0.DBW0, 1 s
   "SDC\DB_SDC_EMS_FLAGS\DB_SDC_EMS_FLAGS.EMS[53]" : Int AT %DB0.DBW0, 1 s
   "SDC\DB_SDC_EMS_FLAGS\DB_SDC_EMS_FLAGS.EMS[54]" : Int AT %DB0.DBW0, 1 s
   "SDC\DB_SDC_EMS_FLAGS\DB_SDC_EMS_FLAGS.EMS[55]" : Int AT %DB0.DBW0, 1 s
   "SDC\DB_SDC_EMS_FLAGS\DB_SDC_EMS_FLAGS.EMS[56]" : Int AT %DB0.DBW0, 1 s
   "SDC\DB_SDC_EMS_FLAGS\DB_SDC_EMS_FLAGS.EMS[57]" : Int AT %DB0.DBW0, 1 s
   "SDC\DB_SDC_EMS_FLAGS\DB_SDC_EMS_FLAGS.EMS[58]" : Int AT %DB0.DBW0, 1 s
   "SDC\DB_SDC_EMS_FLAGS\DB_SDC_EMS_FLAGS.EMS[59]" : Int AT %DB0.DBW0, 1 s
   "SDC\DB_SDC_EMS_FLAGS\DB_SDC_EMS_FLAGS.EMS[60]" : Int AT %DB0.DBW0, 1 s
   "SDC\DB_SDC_EMS_FLAGS\DB_SDC_EMS_FLAGS.EMS[61]" : Int AT %DB0.DBW0, 1 s
   "SDC\DB_SDC_EMS_FLAGS\DB_SDC_EMS_FLAGS.EMS[62]" : Int AT %DB0.DBW0, 1 s
   "SDC\DB_SDC_EMS_FLAGS\DB_SDC_EMS_FLAGS.EMS[63]" : Int AT %DB0.DBW0, 1 s
   "SDC\DB_SDC_EMS_FLAGS\DB_SDC_EMS_FLAGS.EMS[64]" : Int AT %DB0.DBW0, 1 s
   "SDC\DB_SDC_EMS_FLAGS\DB_SDC_EMS_FLAGS.EMS[65]" : Int AT %DB0.DBW0, 1 s
   "SDC\DB_SDC_EMS_FLAGS\DB_SDC_EMS_FLAGS.EMS[66]" : Int AT %DB0.DBW0, 1 s
   "SDC\DB_SDC_EMS_FLAGS\DB_SDC_EMS_FLAGS.EMS[67]" : Int AT %DB0.DBW0, 1 s
   "SDC\DB_SDC_EMS_FLAGS\DB_SDC_EMS_FLAGS.EMS[68]" : Int AT %DB0.DBW0, 1 s
   "SDC\DB_SDC_EMS_FLAGS\DB_SDC_EMS_FLAGS.EMS[69]" : Int AT %DB0.DBW0, 1 s
   "SDC\DB_SDC_EMS_FLAGS\DB_SDC_EMS_FLAGS.EMS[70]" : Int AT %DB0.DBW0, 1 s
   "SDC\DB_SDC_EMS_FLAGS\DB_SDC_EMS_FLAGS.EMS[71]" : Int AT %DB0.DBW0, 1 s
   "SDC\DB_SDC_EMS_FLAGS\DB_SDC_EMS_FLAGS.EMS[72]" : Int AT %DB0.DBW0, 1 s
   "SDC\DB_SDC_EMS_FLAGS\DB_SDC_EMS_FLAGS.EMS[73]" : Int AT %DB0.DBW0, 1 s
   "SDC\DB_SDC_EMS_FLAGS\DB_SDC_EMS_FLAGS.EMS[74]" : Int AT %DB0.DBW0, 1 s
   "SDC\DB_SDC_EMS_FLAGS\DB_SDC_EMS_FLAGS.EMS[75]" : Int AT %DB0.DBW0, 1 s
   "SDC\DB_SDC_EMS_FLAGS\DB_SDC_EMS_FLAGS.EMS[76]" : Int AT %DB0.DBW0, 1 s
   "SDC\DB_SDC_EMS_FLAGS\DB_SDC_EMS_FLAGS.EMS[77]" : Int AT %DB0.DBW0, 1 s
   "SDC\DB_SDC_EMS_FLAGS\DB_SDC_EMS_FLAGS.EMS[78]" : Int AT %DB0.DBW0, 1 s
   "SDC\DB_SDC_EMS_FLAGS\DB_SDC_EMS_FLAGS.EMS[79]" : Int AT %DB0.DBW0, 1 s
   "SDC\DB_SDC_EMS_FLAGS\DB_SDC_EMS_FLAGS.EMS[80]" : Int AT %DB0.DBW0, 1 s
   "SDC\DB_SDC_EMS_FLAGS\DB_SDC_EMS_FLAGS.EMS[81]" : Int AT %DB0.DBW0, 1 s
   "SDC\DB_SDC_EMS_FLAGS\DB_SDC_EMS_FLAGS.EMS[82]" : Int AT %DB0.DBW0, 1 s
   "SDC\DB_SDC_EMS_FLAGS\DB_SDC_EMS_FLAGS.EMS[83]" : Int AT %DB0.DBW0, 1 s
   "SDC\DB_SDC_EMS_FLAGS\DB_SDC_EMS_FLAGS.EMS[84]" : Int AT %DB0.DBW0, 1 s
   "SDC\DB_SDC_EMS_FLAGS\DB_SDC_EMS_FLAGS.EMS[85]" : Int AT %DB0.DBW0, 1 s
   "SDC\DB_SDC_EMS_FLAGS\DB_SDC_EMS_FLAGS.EMS[86]" : Int AT %DB0.DBW0, 1 s
   "SDC\DB_SDC_EMS_FLAGS\DB_SDC_EMS_FLAGS.EMS[87]" : Int AT %DB0.DBW0, 1 s
   "SDC\DB_SDC_EMS_FLAGS\DB_SDC_EMS_FLAGS.EMS[88]" : Int AT %DB0.DBW0, 1 s
   "SDC\DB_SDC_EMS_FLAGS\DB_SDC_EMS_FLAGS.EMS[89]" : Int AT %DB0.DBW0, 1 s
   "SDC\DB_SDC_EMS_FLAGS\DB_SDC_EMS_FLAGS.EMS[90]" : Int AT %DB0.DBW0, 1 s
   "SDC\DB_SDC_EMS_FLAGS\DB_SDC_EMS_FLAGS.EMS[91]" : Int AT %DB0.DBW0, 1 s
   "SDC\DB_SDC_EMS_FLAGS\DB_SDC_EMS_FLAGS.EMS[92]" : Int AT %DB0.DBW0, 1 s
   "SDC\DB_SDC_EMS_FLAGS\DB_SDC_EMS_FLAGS.EMS[93]" : Int AT %DB0.DBW0, 1 s
   "SDC\DB_SDC_EMS_FLAGS\DB_SDC_EMS_FLAGS.EMS[94]" : Int AT %DB0.DBW0, 1 s
   "SDC\DB_SDC_EMS_FLAGS\DB_SDC_EMS_FLAGS.EMS[95]" : Int AT %DB0.DBW0, 1 s
   "SDC\DB_SDC_EMS_FLAGS\DB_SDC_EMS_FLAGS.EMS[96]" : Int AT %DB0.DBW0, 1 s
   "SDC\DB_SDC_EMS_FLAGS\DB_SDC_EMS_FLAGS.EMS[97]" : Int AT %DB0.DBW0, 1 s
   "SDC\DB_SDC_EMS_FLAGS\DB_SDC_EMS_FLAGS.EMS[98]" : Int AT %DB0.DBW0, 1 s